// TIA Portal project "Process visualization with HMI" (V15.1)

(* hardware
DEVICE "S71500/ET200MP station_1"  S7-1500 station
   slot 0: "Rail_0"  Rack  6ES7 590-1***0-0AA0
   slot 0: "PM 190W 120/230VAC"  PM 190W 120/230VAC  6EP1333-4BA00
   slot 1: "PLC_1"  CPU 1516-3 PN/DP  6ES7 516-3AN01-0AB0  V2.6
      slot 3: "CPU display_1"  6ES7591-1BA00-0AA0
   slot 2: "DQ 32x24VDC/0.5A HF_1"  DQ 32x24VDC/0.5A HF  6ES7 522-1BL01-0AB0  V1.1
   slot 3: "DI 32x24VDC HF_1"  DI 32x24VDC HF  6ES7 521-1BL00-0AB0  V2.1
   slot 4: "AQ 4xU/I ST_1"  AQ 4xU/I ST  6ES7 532-5HD00-0AB0  V2.2
   slot 5: "AI 8xU/I/RTD/TC ST_1"  AI 8xU/I/RTD/TC ST  6ES7 531-7KF00-0AB0  V2.2
DEVICE "HMI_1"  TP700 Comfort
   slot 0: "HMI_1"  TP700 Comfort  6AV2 124-0GC01-0AX0  15.1.0.0
   slot 1: "HMI_RT_1"  TP700 Comfort  6AV2 124-0GC01-0AX0  15.1.0.0
   slot 5: "HMI_1.IE_CP_1"  PROFINET Interface  15.0.1.0
      slot 1: "PROFINET Interface_1"  PROFINET Interface
         slot 1: "Port_1"  Port
         slot 2: "Port_2"  Port
   slot 7: "HMI_1.MPI/DP_CP_1"  MPI/DP Interface  15.0.1.0
*)

// ===== PLC "PLC_1"  CPU 1516-3 PN/DP =====

VAR_GLOBAL   // PLC tag table "Full_Tag_Table"
   "Panel Emergency Stop" AT %I2.7 : Bool;
   "Start switch" AT %I0.2 : Bool;
   "Stop switch" AT %I0.3 : Bool;
   "Sort area IR" AT %I0.4 : Bool;
   "Sort Area Inductive" AT %I0.5 : Bool;
   "Sort Solenoid Sensor" AT %I0.6 : Bool;
   "Assembly Chute IR" AT %I0.7 : Bool;
   "Assembly Area Through Beam" AT %I1.1 : Bool;
   "Assembly Area Capacitor" AT %I1.2 : Bool;
   "Assembly Area Inductive" AT %I1.3 : Bool;
   "Reject Area IR" AT %I1.4 : Bool;
   "Reject Solenoid Sensor" AT %I1.5 : Bool;
   "Oven Through Beam" AT %I1.6 : Bool;
   "Loading Area Inductive" AT %I1.7 : Bool;
   "Chain Conveyor" AT %Q0.0 : Bool;
   "Sort Solenoid" AT %Q0.1 : Bool;
   "Reject Solenoid" AT %Q0.2 : Bool;
   "Rotary Solenoid" AT %Q0.3 : Bool;
   "Belt Conveyor Direction" AT %Q0.4 : Bool;
   "System Run_Green Lamp" AT %Q3.0 : Bool;
   "Sysyem Stop_Red Lamp" AT %Q3.2 : Bool;
   "Emergency stop" AT %I1.0 : Bool;
   "Ring Queue counter Full" AT %M4.0 : Bool;
   "Sort Solenoid error" AT %M4.3 : Bool;
   "Counter value" AT %MW0 : Int;
   "Reject Solenoid Error" AT %M4.7 : Bool;
   "HMI_Start" AT %M4.1 : Bool;
   "HMI_Stop" AT %M4.2 : Bool;
   "Counter Reset" AT %M4.4 : Bool;
   "DO_card" AT %QD0 : DWord;
   "DI_card" AT %ID0 : DWord;
   "Assembled part counter value" AT %MW4 : Int;
   "HMI_Emergency" AT %M4.5 : Bool;
   "Output metal peg counter value" AT %MW5 : Int;
   "Output plastic ring counter value" AT %MW6 : Int;
   "Input metal peg counter value" AT %MW8 : Int;
   "Input plastic ring counter value" AT %MW10 : Int;
END_VAR

DATA_BLOCK "Conveyors_AUTOMATIC_DB"   // DB1
{ S7_Optimized_Access := 'TRUE' }
VERSION : 0.1
// stored: InstanceOfName Conveyors_AUTOMATIC
"Conveyors_AUTOMATIC"
BEGIN
END_DATA_BLOCK

DATA_BLOCK "Sort Solenoid active_DB"   // DB2
{ S7_Optimized_Access := 'TRUE' }
VERSION : 0.1
// stored: InstanceOfName Sort Solenoid active
"Sort Solenoid active"
BEGIN
END_DATA_BLOCK

DATA_BLOCK "Sort Solenoid active_DB_1"   // DB3
{ S7_Optimized_Access := 'TRUE' }
VERSION : 0.1
// stored: InstanceOfName Sort Solenoid active
"Sort Solenoid active"
BEGIN
END_DATA_BLOCK

DATA_BLOCK "Solenoid Error_DB"   // DB4
{ S7_Optimized_Access := 'TRUE' }
VERSION : 0.1
// stored: InstanceOfName Solenoid Error
"Solenoid Error"
BEGIN
END_DATA_BLOCK

DATA_BLOCK "Counting_DB"   // DB5
{ S7_Optimized_Access := 'TRUE' }
VERSION : 0.1
// stored: InstanceOfName Counter
"Counter"
BEGIN
END_DATA_BLOCK

DATA_BLOCK "Rotary Solenoid1_DB"   // DB6
{ S7_Optimized_Access := 'TRUE' }
VERSION : 0.1
// stored: InstanceOfName Rotary Solenoid1
"Rotary Solenoid1"
BEGIN
END_DATA_BLOCK

DATA_BLOCK "Component Queue Handling_DB"   // DB7
{ S7_Optimized_Access := 'TRUE' }
VERSION : 0.1
// stored: InstanceOfName Component Queue Handling
"Component Queue Handling"
BEGIN
END_DATA_BLOCK

DATA_BLOCK "Solenoid Error_DB_1"   // DB8
{ S7_Optimized_Access := 'TRUE' }
VERSION : 0.1
// stored: InstanceOfName Solenoid Error
"Solenoid Error"
BEGIN
END_DATA_BLOCK

DATA_BLOCK "Assembled part counter_DB"   // DB9
{ S7_Optimized_Access := 'TRUE' }
VERSION : 0.1
// stored: InstanceOfName Assembled part counter
"Assembled part counter"
BEGIN
END_DATA_BLOCK

DATA_BLOCK "Metal peg after assembly counter_DB"   // DB10
{ S7_Optimized_Access := 'TRUE' }
VERSION : 0.1
// stored: InstanceOfName Output metal peg counter
"Output metal peg counter"
BEGIN
END_DATA_BLOCK

DATA_BLOCK "Plastic ring after assembly counter_DB"   // DB11
{ S7_Optimized_Access := 'TRUE' }
VERSION : 0.1
// stored: InstanceOfName Output plastic ring counter
"Output plastic ring counter"
BEGIN
END_DATA_BLOCK

DATA_BLOCK "Input metal peg counter_DB"   // DB12
{ S7_Optimized_Access := 'TRUE' }
VERSION : 0.1
// stored: InstanceOfName Input metal peg counter
"Input metal peg counter"
BEGIN
END_DATA_BLOCK

DATA_BLOCK "Input plastic ring counter_DB"   // DB13
{ S7_Optimized_Access := 'TRUE' }
VERSION : 0.1
// stored: InstanceOfName Input plastic ring counter
"Input plastic ring counter"
BEGIN
END_DATA_BLOCK

FUNCTION_BLOCK "Conveyors_AUTOMATIC"   // FB1, LAD
TITLE = Conveyors Automatic
{ S7_Optimized_Access := 'TRUE' }
VERSION : 0.1
   VAR_INPUT
      "Start Switch" : Bool;
      "Stop Switch" : Bool;
      "Emergency Stop" : Bool;
      "Sort Solenoid Error" : Bool;
      "Panel Emergency Stop" : Bool;
      "Reject Solenoid Error" : Bool;
      H_Start : Bool;
      H_Stop : Bool;
      H_Emergency : Bool;
   END_VAR
   VAR_OUTPUT
      "Chain Conveyor" : Bool;
      "Belt Conveyor" : Bool;
      "System Enable_OK" : Bool;
      "System Enable_not_OK" : Bool;
   END_VAR
   VAR
      Memory_Automatic_Start_Stop : Bool;
   END_VAR
BEGIN

REGION Network 1: System Enable_OK and Conveyor Run
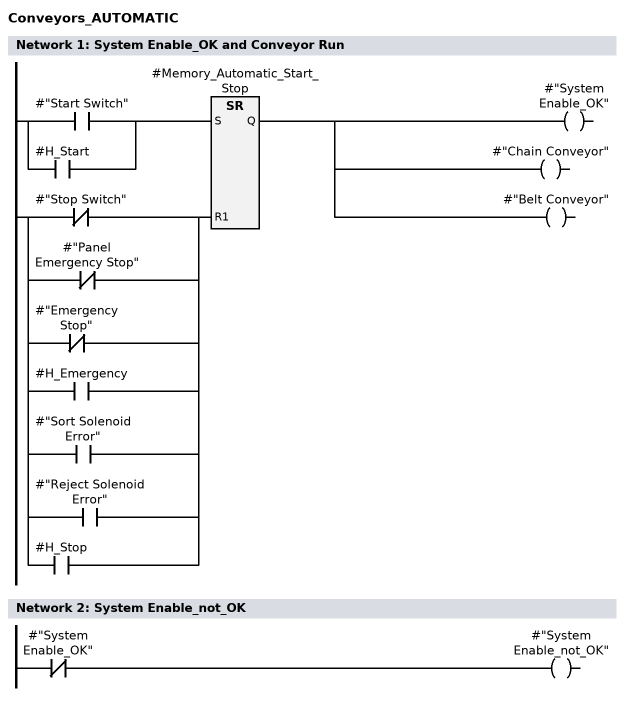
   RUNG wire#powerrail
      Contact( #"Start Switch" )
      wire#w1
      S_SR(operand := #Memory_Automatic_Start_Stop, r1 := wire#w2)
      wire#w3
      Coil( #"System Enable_OK" )
   END_RUNG
   RUNG wire#powerrail
      Contact( #H_Start )
   END_RUNG wire#w1
   RUNG wire#powerrail
      I_Contact( #"Stop Switch" )
   END_RUNG wire#w2
   RUNG wire#powerrail
      I_Contact( #"Panel Emergency Stop" )
   END_RUNG wire#w2
   RUNG wire#powerrail
      I_Contact( #"Emergency Stop" )
   END_RUNG wire#w2
   RUNG wire#powerrail
      Contact( #H_Emergency )
   END_RUNG wire#w2
   RUNG wire#powerrail
      Contact( #"Sort Solenoid Error" )
   END_RUNG wire#w2
   RUNG wire#powerrail
      Contact( #"Reject Solenoid Error" )
   END_RUNG wire#w2
   RUNG wire#powerrail
      Contact( #H_Stop )
   END_RUNG wire#w2
   RUNG wire#w3
      Coil( #"Chain Conveyor" )
   END_RUNG
   RUNG wire#w3
      Coil( #"Belt Conveyor" )
   END_RUNG
   // the same network as SCL:
   IF #"Start Switch" OR #H_Start THEN
       #Memory_Automatic_Start_Stop := TRUE;   // SR flip-flop
   END_IF;
   IF NOT #"Stop Switch" OR NOT #"Panel Emergency Stop" OR NOT #"Emergency Stop" OR #H_Emergency OR #"Sort Solenoid Error" OR #"Reject Solenoid Error" OR #H_Stop THEN
       #Memory_Automatic_Start_Stop := FALSE;
   END_IF;
   #"System Enable_OK" := #Memory_Automatic_Start_Stop;
   #"Chain Conveyor" := #Memory_Automatic_Start_Stop;
   #"Belt Conveyor" := #Memory_Automatic_Start_Stop;
END_REGION

REGION Network 2: System Enable_not_OK
   RUNG wire#powerrail
      I_Contact( #"System Enable_OK" )
      Coil( #"System Enable_not_OK" )
   END_RUNG
   // the same network as SCL:
   #"System Enable_not_OK" := NOT #"System Enable_OK";
END_REGION
END_FUNCTION_BLOCK

FUNCTION_BLOCK "Sort Solenoid active"   // FB2, LAD
TITLE = Sort Solenoid active
{ S7_Optimized_Access := 'TRUE' }
VERSION : 0.1
   VAR_INPUT
      "Sort Area IR" : Bool;
      "Sort Area Inductive" : Bool;
      "Ring Queue counter full" : Bool;
   END_VAR
   VAR_OUTPUT
      "Sort Solenoid" : Bool;
   END_VAR
   VAR
      "Component Pass Delay" : Bool;
      "SR_Sort solenoid on Timer" : Bool;
      "SR_Component pass Delay" : Bool;
      IEC_Timer_0_Instance : TON_TIME;
      IEC_Timer_0_Instance_1 : TON_TIME;
   END_VAR
BEGIN

REGION Network 1: Sort Solenoid activate in case of plastic ring presence
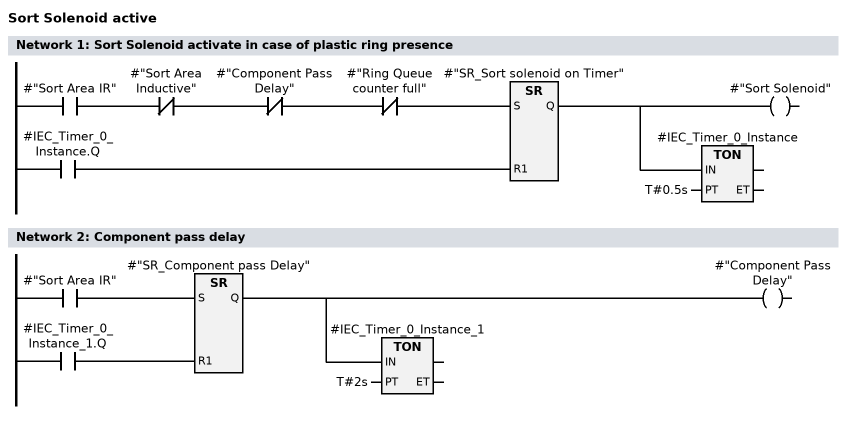
   IF #"Sort Area IR" AND NOT #"Sort Area Inductive" AND NOT #"Component Pass Delay" AND NOT #"Ring Queue counter full" THEN
       #"SR_Sort solenoid on Timer" := TRUE;   // SR flip-flop
   END_IF;
   IF #IEC_Timer_0_Instance.Q THEN #"SR_Sort solenoid on Timer" := FALSE; END_IF;
   #"Sort Solenoid" := #"SR_Sort solenoid on Timer";
   #IEC_Timer_0_Instance(IN := #"SR_Sort solenoid on Timer", PT := T#0.5s);   // TON
END_REGION

REGION Network 2: Component pass delay
   IF #"Sort Area IR" THEN
       #"SR_Component pass Delay" := TRUE;   // SR flip-flop
   END_IF;
   IF #IEC_Timer_0_Instance_1.Q THEN #"SR_Component pass Delay" := FALSE; END_IF;
   #"Component Pass Delay" := #"SR_Component pass Delay";
   #IEC_Timer_0_Instance_1(IN := #"SR_Component pass Delay", PT := T#2s);   // TON
END_REGION
END_FUNCTION_BLOCK

FUNCTION_BLOCK "Solenoid Error"   // FB3, LAD
TITLE = Solenoid error
{ S7_Optimized_Access := 'TRUE' }
VERSION : 0.1
   VAR_INPUT
      "Solenoid on" : Bool;
      "Solenoid sensor" : Bool;
   END_VAR
   VAR_OUTPUT
      "Solenoid error" : Bool;
   END_VAR
   VAR
      "Hold off delay" : Bool;
      IEC_Timer_0_Instance : TON_TIME;
   END_VAR
BEGIN

REGION Network 1: Solenoid error
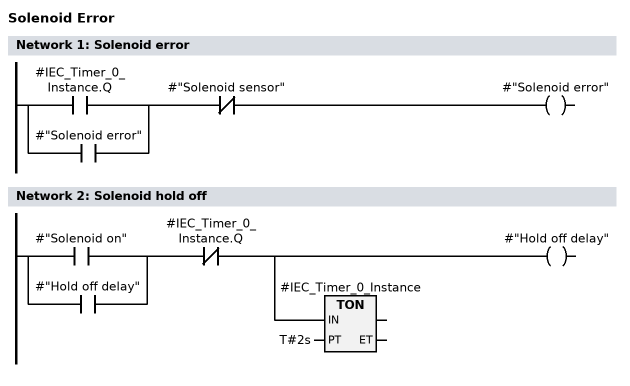
   RUNG wire#powerrail
      Contact( #IEC_Timer_0_Instance.Q )
      wire#w1
      I_Contact( #"Solenoid sensor" )
      Coil( #"Solenoid error" )
   END_RUNG
   RUNG wire#powerrail
      Contact( #"Solenoid error" )
   END_RUNG wire#w1
   // the same network as SCL:
   #"Solenoid error" := (#IEC_Timer_0_Instance.Q OR #"Solenoid error") AND NOT #"Solenoid sensor";
END_REGION

REGION Network 2: Solenoid hold off
   #"Hold off delay" := (#"Solenoid on" OR #"Hold off delay") AND NOT #IEC_Timer_0_Instance.Q;
   #IEC_Timer_0_Instance(IN := #"Hold off delay", PT := T#2s);   // TON
END_REGION
END_FUNCTION_BLOCK

FUNCTION_BLOCK "Counter"   // FB4, LAD
{ S7_Optimized_Access := 'TRUE' }
VERSION : 0.1
   VAR_INPUT
      "Sort Solenoid" : Bool;
      "Rotary Solenoid" : Bool;
      "Reset counter" : Bool;
   END_VAR
   VAR_OUTPUT
      "Counter value" : Int;
      "Ring Queue counter full" : Bool;
   END_VAR
   VAR RETAIN
      IEC_Counter_0_Instance : CTUD_INT;
   END_VAR
BEGIN

REGION Network 1
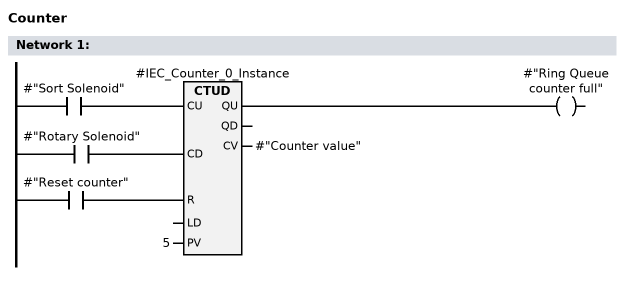
   #IEC_Counter_0_Instance(CU := #"Sort Solenoid",   // CTUD
                           CD := #"Rotary Solenoid",
                           R := #"Reset counter",
                           PV := 5,
                           CV => #"Counter value");
   #"Ring Queue counter full" := #IEC_Counter_0_Instance.QU;
END_REGION
END_FUNCTION_BLOCK

FUNCTION_BLOCK "Rotary Solenoid1"   // FB5, LAD
{ S7_Optimized_Access := 'TRUE' }
VERSION : 0.1
   VAR_INPUT
      "Assembly chute IR" : Bool;
      "Counter value" : Int;
   END_VAR
   VAR_OUTPUT
      "Rotary Solenoid" : Bool;
   END_VAR
   VAR
      "Rotary Solenoid on Timer" : Bool;
      IEC_Timer_0_Instance : TON_TIME;
      "Component pass delay" : Bool;
      "SR_Component pass delay" : Bool;
      IEC_Timer_0_Instance_2 : TON_TIME;
      IEC_Timer_0_Instance_1 : TON_TIME;
   END_VAR
BEGIN

REGION Network 1: Rotary Solenoid
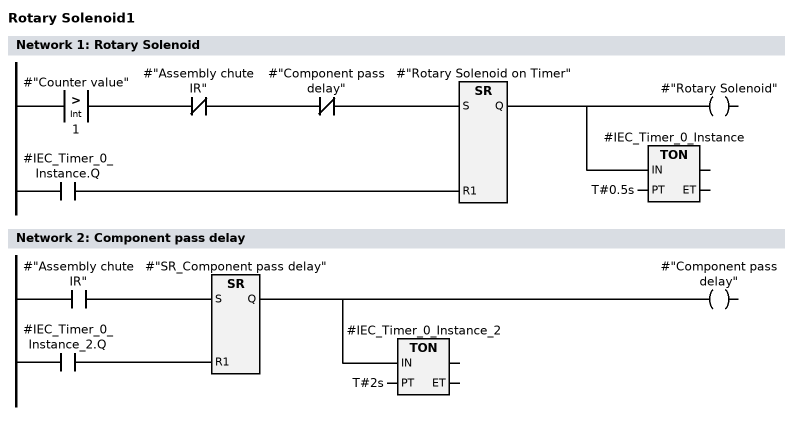
   IF (#"Counter value" > 1) AND NOT #"Assembly chute IR" AND NOT #"Component pass delay" THEN
       #"Rotary Solenoid on Timer" := TRUE;   // SR flip-flop
   END_IF;
   IF #IEC_Timer_0_Instance.Q THEN #"Rotary Solenoid on Timer" := FALSE; END_IF;
   #"Rotary Solenoid" := #"Rotary Solenoid on Timer";
   #IEC_Timer_0_Instance(IN := #"Rotary Solenoid on Timer", PT := T#0.5s);   // TON
END_REGION

REGION Network 2: Component pass delay
   IF #"Assembly chute IR" THEN
       #"SR_Component pass delay" := TRUE;   // SR flip-flop
   END_IF;
   IF #IEC_Timer_0_Instance_2.Q THEN #"SR_Component pass delay" := FALSE; END_IF;
   #"Component pass delay" := #"SR_Component pass delay";
   #IEC_Timer_0_Instance_2(IN := #"SR_Component pass delay", PT := T#2s);   // TON
END_REGION
END_FUNCTION_BLOCK

FUNCTION_BLOCK "Component Queue Handling"   // FB6, LAD
TITLE = Component Queue Handling
{ S7_Optimized_Access := 'TRUE' }
VERSION : 0.1
   VAR_INPUT
      "Start Switch" : Bool;
      "Assembly Area Capacitive" : Bool;
      "Assembly Area Inductive" : Bool;
      "Reject Area IR" : Bool;
      "Assembly Area Through Beam" : Bool;
   END_VAR
   VAR_OUTPUT
      "Reject Solenoid" : Bool;
   END_VAR
   VAR
      "Assembly Complete" : Bool;
      "Pointer Register" : Word;
      "Data Register" : Word;
      "SHL Memory" : Bool;
      "SHR Memory" : Bool;
      "And Result" : Word;
      SR_Reject : Bool;
      IEC_Timer_0_Instance : TON_TIME;
   END_VAR
   VAR_TEMP   // added for the SCL form of the ladder/FBD networks
      _w1 : Bool;
   END_VAR
BEGIN

REGION Network 1: data and pointer register
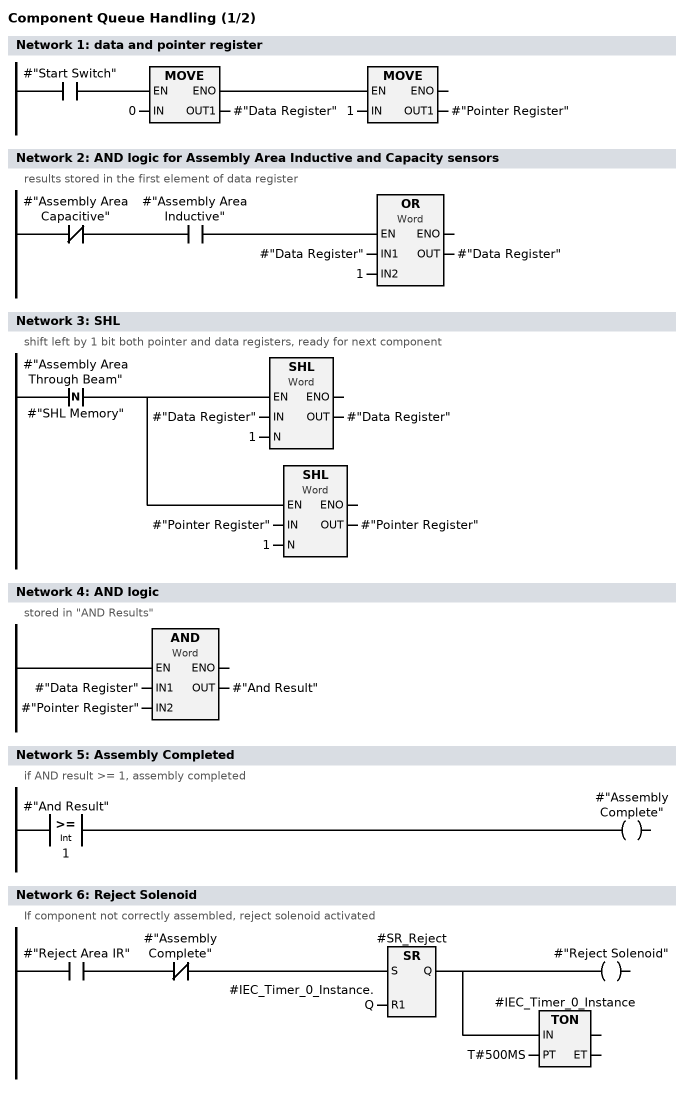
   RUNG wire#powerrail
      Contact( #"Start Switch" )
      Move(in := 0, out1 => #"Data Register")
      Move(in := 1, out1 => #"Pointer Register")
   END_RUNG
   // the same network as SCL:
   IF #"Start Switch" THEN
       #"Data Register" := 0;
       #"Pointer Register" := 1;
   END_IF;
END_REGION

REGION Network 2: AND logic for Assembly Area Inductive and Capacity sensors
   // results stored in the first element of data register
   IF NOT #"Assembly Area Capacitive" AND #"Assembly Area Inductive" THEN
       #"Data Register" := #"Data Register" OR 1;
   END_IF;
END_REGION

REGION Network 3: SHL
   // shift left by 1 bit both pointer and data registers, ready for next component
   RUNG wire#powerrail
      N_Contact(operand := #"Assembly Area Through Beam", bit := #"SHL Memory")
      wire#w1
      { S7_Templates := "SrcType := Word" } Shl(in := #"Data Register", n := 1, out => #"Data Register")
   END_RUNG
   RUNG wire#w1
      { S7_Templates := "SrcType := Word" } Shl(in := #"Pointer Register", n := 1, out => #"Pointer Register")
   END_RUNG
   // the same network as SCL:
   #_w1 := NOT #"Assembly Area Through Beam" AND #"SHL Memory";   // falling edge of #"Assembly Area Through Beam"
   #"SHL Memory" := #"Assembly Area Through Beam";
   IF #_w1 THEN
       #"Data Register" := SHL(IN := #"Data Register", N := 1);
       #"Pointer Register" := SHL(IN := #"Pointer Register", N := 1);
   END_IF;
END_REGION

REGION Network 4: AND logic
   // stored in "AND Results"
   RUNG wire#powerrail
      { S7_Templates := "SrcType := Word" } And(in1 := #"Data Register", in2 := #"Pointer Register", out => #"And Result")
   END_RUNG
   // the same network as SCL:
   #"And Result" := #"Data Register" AND #"Pointer Register";
END_REGION

REGION Network 5: Assembly Completed
   // if AND result >= 1, assembly completed
   RUNG wire#powerrail
      { S7_Templates := "SrcType := Int" } GE_Contact(in1 := #"And Result", in2 := 1)
      Coil( #"Assembly Complete" )
   END_RUNG
   // the same network as SCL:
   #"Assembly Complete" := #"And Result" >= 1;
END_REGION

REGION Network 6: Reject Solenoid
   // If component not correctly assembled, reject solenoid activated
   IF #"Reject Area IR" AND NOT #"Assembly Complete" THEN
       #SR_Reject := TRUE;   // SR flip-flop
   END_IF;
   IF #IEC_Timer_0_Instance.Q THEN #SR_Reject := FALSE; END_IF;
   #"Reject Solenoid" := #SR_Reject;
   #IEC_Timer_0_Instance(IN := #SR_Reject, PT := T#500MS);   // TON
END_REGION

REGION Network 7: SHR
   // when component left assembly area, shift right by 1 bit
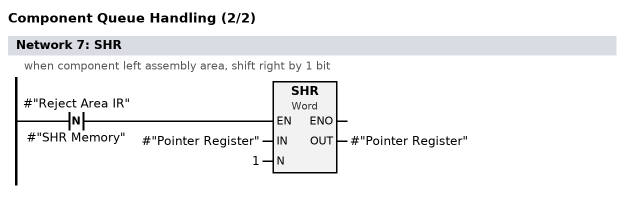
   RUNG wire#powerrail
      N_Contact(operand := #"Reject Area IR", bit := #"SHR Memory")
      { S7_Templates := "SrcType := Word" } Shr(in := #"Pointer Register", n := 1, out => #"Pointer Register")
   END_RUNG
   // the same network as SCL:
   #_w1 := NOT #"Reject Area IR" AND #"SHR Memory";   // falling edge of #"Reject Area IR"
   #"SHR Memory" := #"Reject Area IR";
   IF #_w1 THEN #"Pointer Register" := SHR(IN := #"Pointer Register", N := 1); END_IF;
END_REGION
END_FUNCTION_BLOCK

FUNCTION_BLOCK "Assembled part counter"   // FB7, LAD
TITLE = Assembled part counter
{ S7_Optimized_Access := 'TRUE' }
VERSION : 0.1
   VAR_INPUT
      "Reject area IR" : Bool;
      "Reject solenoid" : Bool;
      "Reset counter" : Bool;
   END_VAR
   VAR_OUTPUT
      "Assembled part counter value" : Int;
   END_VAR
   VAR RETAIN
      IEC_Counter_0_Instance : CTU_INT;
   END_VAR
BEGIN

REGION Network 1: Counter for assembled parts
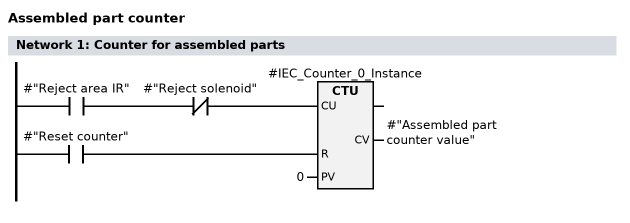
   #IEC_Counter_0_Instance(CU := #"Reject area IR" AND NOT #"Reject solenoid",   // CTU
                           R := #"Reset counter",
                           PV := 0,
                           CV => #"Assembled part counter value");
END_REGION
END_FUNCTION_BLOCK

FUNCTION_BLOCK "Output metal peg counter"   // FB8, LAD
{ S7_Optimized_Access := 'TRUE' }
VERSION : 0.1
   VAR_INPUT
      "Assembly Area Inductive" : Bool;
      "Assembly Area Capacitive" : Bool;
      "Assembly Area thru beam" : Bool;
      "Reset counter" : Bool;
   END_VAR
   VAR_OUTPUT
      "Metal peg" : Int;
   END_VAR
   VAR RETAIN
      IEC_Counter_0_Instance : CTU_INT;
   END_VAR
BEGIN

REGION Network 1: Metal peg counter
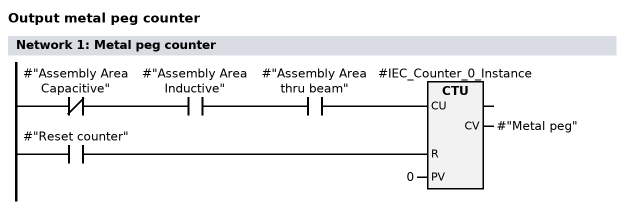
   #IEC_Counter_0_Instance(CU := NOT #"Assembly Area Capacitive" AND #"Assembly Area Inductive" AND #"Assembly Area thru beam",   // CTU
                           R := #"Reset counter",
                           PV := 0,
                           CV => #"Metal peg");
END_REGION
END_FUNCTION_BLOCK

FUNCTION_BLOCK "Output plastic ring counter"   // FB9, LAD
{ S7_Optimized_Access := 'TRUE' }
VERSION : 0.1
   VAR_INPUT
      "Assembly Area Inductive" : Bool;
      "Assembly Area Capacitive" : Bool;
      "Assembly Area thru beam" : Bool;
      "Reset counter" : Bool;
   END_VAR
   VAR_OUTPUT
      "Plastic ring" : Int;
   END_VAR
   VAR RETAIN
      IEC_Counter_0_Instance : CTU_INT;
   END_VAR
BEGIN

REGION Network 1: Plastic ring counter
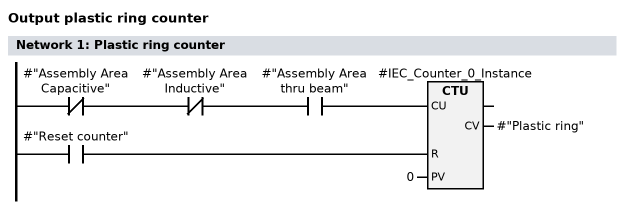
   #IEC_Counter_0_Instance(CU := NOT #"Assembly Area Capacitive" AND NOT #"Assembly Area Inductive" AND #"Assembly Area thru beam",   // CTU
                           R := #"Reset counter",
                           PV := 0,
                           CV => #"Plastic ring");
END_REGION
END_FUNCTION_BLOCK

FUNCTION_BLOCK "Input metal peg counter"   // FB10, LAD
{ S7_Optimized_Access := 'TRUE' }
VERSION : 0.1
   VAR_INPUT
      "Sort Area IR" : Bool;
      "Sort Area inductive" : Bool;
      "Reset counter" : Bool;
   END_VAR
   VAR_OUTPUT
      "Input metal peg" : Int;
   END_VAR
   VAR RETAIN
      IEC_Counter_0_Instance : CTU_INT;
   END_VAR
BEGIN

REGION Network 1: Input Metal Peg counter
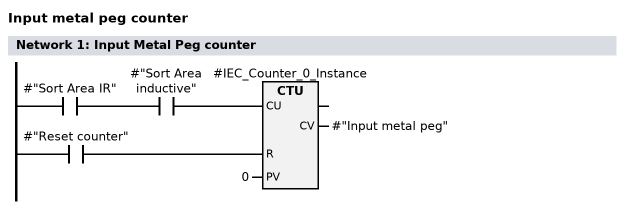
   #IEC_Counter_0_Instance(CU := #"Sort Area IR" AND #"Sort Area inductive",   // CTU
                           R := #"Reset counter",
                           PV := 0,
                           CV => #"Input metal peg");
END_REGION
END_FUNCTION_BLOCK

FUNCTION_BLOCK "Input plastic ring counter"   // FB11, LAD
{ S7_Optimized_Access := 'TRUE' }
VERSION : 0.1
   VAR_INPUT
      "Sort Area IR" : Bool;
      "Sort Area inductive" : Bool;
      "Reset counter" : Bool;
   END_VAR
   VAR_OUTPUT
      "Input plastic ring" : Int;
   END_VAR
   VAR RETAIN
      IEC_Counter_0_Instance : CTU_INT;
   END_VAR
BEGIN

REGION Network 1: Input plastic ring counter
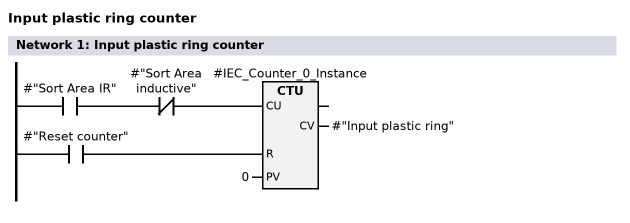
   #IEC_Counter_0_Instance(CU := #"Sort Area IR" AND NOT #"Sort Area inductive",   // CTU
                           R := #"Reset counter",
                           PV := 0,
                           CV => #"Input plastic ring");
END_REGION
END_FUNCTION_BLOCK

ORGANIZATION_BLOCK "Main"   // OB1, LAD, ProgramCycle
TITLE = "Main Program Sweep (Cycle)"
{ S7_Optimized_Access := 'TRUE' }
VERSION : 0.1
   VAR_INPUT
      Initial_Call : Bool;   // Initial call of this OB
      Remanence : Bool;   // =True, if remanent data are available
   END_VAR
BEGIN

REGION Network 1: System Run OK and conveyors start
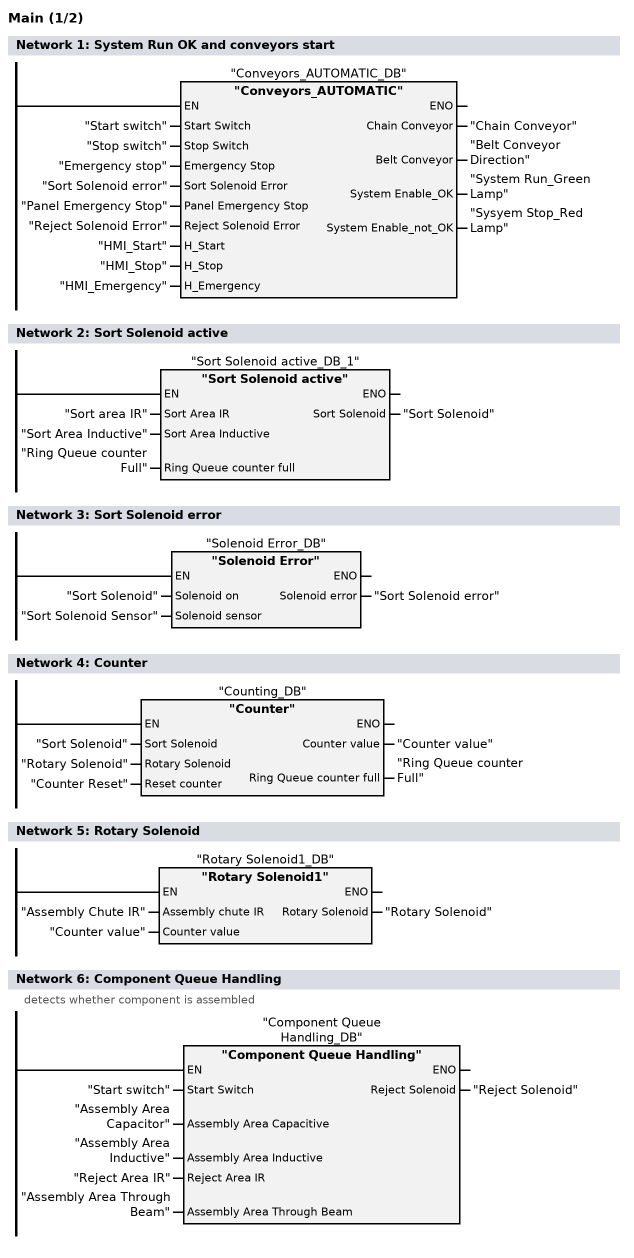
   RUNG wire#powerrail
      "Conveyors_AUTOMATIC_DB"("Start Switch" := "Start switch", "Stop Switch" := "Stop switch", "Emergency Stop" := "Emergency stop", "Sort Solenoid Error" := "Sort Solenoid error", "Panel Emergency Stop" := "Panel Emergency Stop", "Reject Solenoid Error" := "Reject Solenoid Error", H_Start := "HMI_Start", H_Stop := "HMI_Stop", H_Emergency := "HMI_Emergency", "Chain Conveyor" => "Chain Conveyor", "Belt Conveyor" => "Belt Conveyor Direction", "System Enable_OK" => "System Run_Green Lamp", "System Enable_not_OK" => "Sysyem Stop_Red Lamp")
   END_RUNG
   // the same network as SCL:
   "Conveyors_AUTOMATIC_DB"("Start Switch" := "Start switch",   // "Conveyors_AUTOMATIC"
                           "Stop Switch" := "Stop switch",
                           "Emergency Stop" := "Emergency stop",
                           "Sort Solenoid Error" := "Sort Solenoid error",
                           "Panel Emergency Stop" := "Panel Emergency Stop",
                           "Reject Solenoid Error" := "Reject Solenoid Error",
                           H_Start := "HMI_Start",
                           H_Stop := "HMI_Stop",
                           H_Emergency := "HMI_Emergency",
                           "Chain Conveyor" => "Chain Conveyor",
                           "Belt Conveyor" => "Belt Conveyor Direction",
                           "System Enable_OK" => "System Run_Green Lamp",
                           "System Enable_not_OK" => "Sysyem Stop_Red Lamp");
END_REGION

REGION Network 2: Sort Solenoid active
   RUNG wire#powerrail
      "Sort Solenoid active_DB_1"("Sort Area IR" := "Sort area IR", "Sort Area Inductive" := "Sort Area Inductive", "Ring Queue counter full" := "Ring Queue counter Full", "Sort Solenoid" => "Sort Solenoid")
   END_RUNG
   // the same network as SCL:
   "Sort Solenoid active_DB_1"("Sort Area IR" := "Sort area IR",   // "Sort Solenoid active"
                           "Sort Area Inductive" := "Sort Area Inductive",
                           "Ring Queue counter full" := "Ring Queue counter Full",
                           "Sort Solenoid" => "Sort Solenoid");
END_REGION

REGION Network 3: Sort Solenoid error
   RUNG wire#powerrail
      "Solenoid Error_DB"("Solenoid on" := "Sort Solenoid", "Solenoid sensor" := "Sort Solenoid Sensor", "Solenoid error" => "Sort Solenoid error")
   END_RUNG
   // the same network as SCL:
   "Solenoid Error_DB"("Solenoid on" := "Sort Solenoid",   // "Solenoid Error"
                       "Solenoid sensor" := "Sort Solenoid Sensor",
                       "Solenoid error" => "Sort Solenoid error");
END_REGION

REGION Network 4: Counter
   RUNG wire#powerrail
      "Counting_DB"("Sort Solenoid" := "Sort Solenoid", "Rotary Solenoid" := "Rotary Solenoid", "Reset counter" := "Counter Reset", "Counter value" => "Counter value", "Ring Queue counter full" => "Ring Queue counter Full")
   END_RUNG
   // the same network as SCL:
   "Counting_DB"("Sort Solenoid" := "Sort Solenoid",   // "Counter"
                 "Rotary Solenoid" := "Rotary Solenoid",
                 "Reset counter" := "Counter Reset",
                 "Counter value" => "Counter value",
                 "Ring Queue counter full" => "Ring Queue counter Full");
END_REGION

REGION Network 5: Rotary Solenoid
   RUNG wire#powerrail
      "Rotary Solenoid1_DB"("Assembly chute IR" := "Assembly Chute IR", "Counter value" := "Counter value", "Rotary Solenoid" => "Rotary Solenoid")
   END_RUNG
   // the same network as SCL:
   "Rotary Solenoid1_DB"("Assembly chute IR" := "Assembly Chute IR",   // "Rotary Solenoid1"
                         "Counter value" := "Counter value",
                         "Rotary Solenoid" => "Rotary Solenoid");
END_REGION

REGION Network 6: Component Queue Handling
   // detects whether component is assembled
   RUNG wire#powerrail
      "Component Queue Handling_DB"("Start Switch" := "Start switch", "Assembly Area Capacitive" := "Assembly Area Capacitor", "Assembly Area Inductive" := "Assembly Area Inductive", "Reject Area IR" := "Reject Area IR", "Assembly Area Through Beam" := "Assembly Area Through Beam", "Reject Solenoid" => "Reject Solenoid")
   END_RUNG
   // the same network as SCL:
   "Component Queue Handling_DB"("Start Switch" := "Start switch",   // "Component Queue Handling"
                           "Assembly Area Capacitive" := "Assembly Area Capacitor",
                           "Assembly Area Inductive" := "Assembly Area Inductive",
                           "Reject Area IR" := "Reject Area IR",
                           "Assembly Area Through Beam" := "Assembly Area Through Beam",
                           "Reject Solenoid" => "Reject Solenoid");
END_REGION

REGION Network 7: Reject Solenoid error
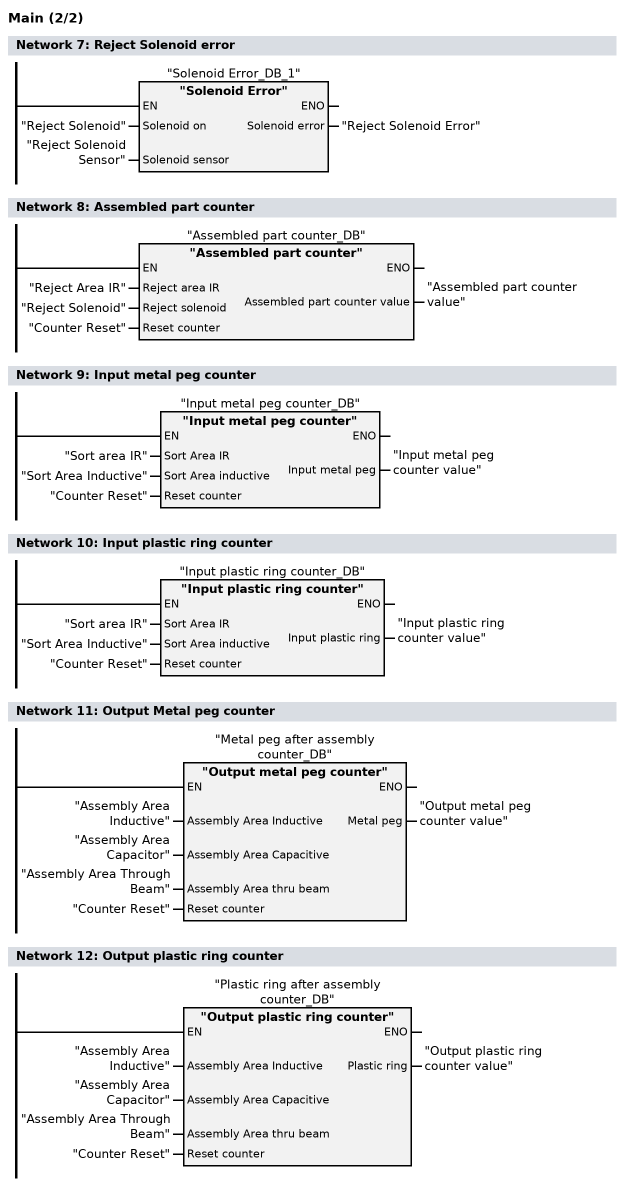
   RUNG wire#powerrail
      "Solenoid Error_DB_1"("Solenoid on" := "Reject Solenoid", "Solenoid sensor" := "Reject Solenoid Sensor", "Solenoid error" => "Reject Solenoid Error")
   END_RUNG
   // the same network as SCL:
   "Solenoid Error_DB_1"("Solenoid on" := "Reject Solenoid",   // "Solenoid Error"
                         "Solenoid sensor" := "Reject Solenoid Sensor",
                         "Solenoid error" => "Reject Solenoid Error");
END_REGION

REGION Network 8: Assembled part counter
   RUNG wire#powerrail
      "Assembled part counter_DB"("Reject area IR" := "Reject Area IR", "Reject solenoid" := "Reject Solenoid", "Reset counter" := "Counter Reset", "Assembled part counter value" => "Assembled part counter value")
   END_RUNG
   // the same network as SCL:
   "Assembled part counter_DB"("Reject area IR" := "Reject Area IR",   // "Assembled part counter"
                           "Reject solenoid" := "Reject Solenoid",
                           "Reset counter" := "Counter Reset",
                           "Assembled part counter value" => "Assembled part counter value");
END_REGION

REGION Network 9: Input metal peg counter
   RUNG wire#powerrail
      "Input metal peg counter_DB"("Sort Area IR" := "Sort area IR", "Sort Area inductive" := "Sort Area Inductive", "Reset counter" := "Counter Reset", "Input metal peg" => "Input metal peg counter value")
   END_RUNG
   // the same network as SCL:
   "Input metal peg counter_DB"("Sort Area IR" := "Sort area IR",   // "Input metal peg counter"
                           "Sort Area inductive" := "Sort Area Inductive",
                           "Reset counter" := "Counter Reset",
                           "Input metal peg" => "Input metal peg counter value");
END_REGION

REGION Network 10: Input plastic ring counter
   RUNG wire#powerrail
      "Input plastic ring counter_DB"("Sort Area IR" := "Sort area IR", "Sort Area inductive" := "Sort Area Inductive", "Reset counter" := "Counter Reset", "Input plastic ring" => "Input plastic ring counter value")
   END_RUNG
   // the same network as SCL:
   "Input plastic ring counter_DB"("Sort Area IR" := "Sort area IR",   // "Input plastic ring counter"
                           "Sort Area inductive" := "Sort Area Inductive",
                           "Reset counter" := "Counter Reset",
                           "Input plastic ring" => "Input plastic ring counter value");
END_REGION

REGION Network 11: Output Metal peg counter
   RUNG wire#powerrail
      "Metal peg after assembly counter_DB"("Assembly Area Inductive" := "Assembly Area Inductive", "Assembly Area Capacitive" := "Assembly Area Capacitor", "Assembly Area thru beam" := "Assembly Area Through Beam", "Reset counter" := "Counter Reset", "Metal peg" => "Output metal peg counter value")
   END_RUNG
   // the same network as SCL:
   "Metal peg after assembly counter_DB"("Assembly Area Inductive" := "Assembly Area Inductive",   // "Output metal peg counter"
                           "Assembly Area Capacitive" := "Assembly Area Capacitor",
                           "Assembly Area thru beam" := "Assembly Area Through Beam",
                           "Reset counter" := "Counter Reset",
                           "Metal peg" => "Output metal peg counter value");
END_REGION

REGION Network 12: Output plastic ring counter
   RUNG wire#powerrail
      "Plastic ring after assembly counter_DB"("Assembly Area Inductive" := "Assembly Area Inductive", "Assembly Area Capacitive" := "Assembly Area Capacitor", "Assembly Area thru beam" := "Assembly Area Through Beam", "Reset counter" := "Counter Reset", "Plastic ring" => "Output plastic ring counter value")
   END_RUNG
   // the same network as SCL:
   "Plastic ring after assembly counter_DB"("Assembly Area Inductive" := "Assembly Area Inductive",   // "Output plastic ring counter"
                           "Assembly Area Capacitive" := "Assembly Area Capacitor",
                           "Assembly Area thru beam" := "Assembly Area Through Beam",
                           "Reset counter" := "Counter Reset",
                           "Plastic ring" => "Output plastic ring counter value");
END_REGION
END_ORGANIZATION_BLOCK

(* ===== HMI "HMI_RT_1" =====
system functions are stored by id; their names below are inferred from use
connection "HMI_Connection_1": ETHERNET, S7_1500_OMS

HMI tags "Default tag table"
   "Counter value" : Int = PLC "Counter value" AT %MW0, 100 ms
   "Sort Solenoid Sensor" : Bool = PLC "Sort Solenoid Sensor" AT %I0.6, 100 ms
   "Ring Queue counter Full" : Bool = PLC "Ring Queue counter Full" AT %M4.0, 100 ms
   "Counter Reset" : Bool = PLC "Counter Reset" AT %M4.4, 100 ms
   "HMI_Stop" : Bool = PLC HMI_Stop AT %M4.2, 100 ms
   "HMI_Start" : Bool = PLC HMI_Start AT %M4.1, 100 ms
   "Emergency stop" : Bool = PLC "Emergency stop" AT %I1.0, 100 ms
   "Stop switch" : Bool = PLC "Stop switch" AT %I0.3, 100 ms
   "System Run_Green Lamp" : Bool = PLC "System Run_Green Lamp" AT %Q3.0, 100 ms
   "Sysyem Stop_Red Lamp" : Bool = PLC "Sysyem Stop_Red Lamp" AT %Q3.2, 100 ms
   "Chain Conveyor" : Bool = PLC "Chain Conveyor" AT %Q0.0, 100 ms
   "Sort area IR" : Bool = PLC "Sort area IR" AT %I0.4, 100 ms
   "Sort Area Inductive" : Bool = PLC "Sort Area Inductive" AT %I0.5, 100 ms
   "Assembly Area Inductive" : Bool = PLC "Assembly Area Inductive" AT %I1.3, 100 ms
   "Assembly Area Capacitor" : Bool = PLC "Assembly Area Capacitor" AT %I1.2, 100 ms
   "Assembly Chute IR" : Bool = PLC "Assembly Chute IR" AT %I0.7, 100 ms
   "Reject Solenoid" : Bool = PLC "Reject Solenoid" AT %Q0.2, 100 ms
   "Reject Solenoid Sensor" : Bool = PLC "Reject Solenoid Sensor" AT %I1.5, 100 ms
   "Belt Conveyor Direction" : Bool = PLC "Belt Conveyor Direction" AT %Q0.4, 100 ms
   "Assembly Area Through Beam" : Bool = PLC "Assembly Area Through Beam" AT %I1.1, 100 ms
   "Assembled part counter value" : Int = PLC "Assembled part counter value" AT %MW4, 100 ms
   "HMI_Emergency" : Bool = PLC HMI_Emergency AT %M4.5, 100 ms
   "Metal peg counter value" : Int = PLC "Output metal peg counter value" AT %MW5, 1 s
   "Plastic ring counter value" : Int = PLC "Output plastic ring counter value" AT %MW6, 1 s
   "Input metal peg counter value" : Int = PLC "Input metal peg counter value" AT %MW8, 1 s
   "Input plastic ring counter value" : Int = PLC "Input plastic ring counter value" AT %MW10, 1 s

Template "Template_1" 800x480
   Button "Exit" at 720,420 size 78x58; TextOff 'Exit'; PictureOff "ExitRuntime_TP700_Comfort_TR"; PictureOn "ExitRuntime_TP700_Comfort_TR"
      on Release: StopRuntime(0)
   Button "Template_Button" at 640,420 size 78x58; TextOff 'Text'
   Button "Template_Button_1" at 560,420 size 78x58; TextOff 'Text'
   Button "Template_Button_2" at 480,420 size 78x58; TextOff 'Text'
   Button "Template_Button_3" at 400,420 size 78x58; TextOff 'Text'
   Button "Template_Button_4" at 321,420 size 78x58; TextOff 'Text'
   Button "Template_Button_5" at 241,420 size 78x58; TextOff 'Text'
   Button "Template_Button_6" at 161,420 size 78x58; TextOff 'Text'
   Button "Template_Button_7" at 81,420 size 78x58; TextOff 'Text'
   Button "Start screen" at 1,420 size 78x58; TextOff 'Start screen'; PictureOff "NavigateHome_TP700_Comfort_TR"; PictureOn "NavigateHome_TP700_Comfort_TR"
      on Release: ActivateScreen("Sorting Station Overview", 0)

screen "Sorting Station Overview" 800x480, template "Template_1"
   TextField "HmiScreenItemData_5" at 80,196 size 640x25; Text 'Welcome to HMI_1 (TP700 Comfort)!'
   Button "HmiScreenItemData" at 36,36 size 159x47; TextOff 'System Control'; PictureOff "Navigates to System Control for TP700 Comfort 15.1.0.0"; PictureOn "Navigates to System Control for TP700 Comfort 15.1.0.0"
      on Release: ActivateScreen("System Control", 0)
   Button "HmiScreenItemData_1" at 36,95 size 159x47; TextOff 'Input/Output'; PictureOff "Navigates to Input/Output for TP700 Comfort 15.1.0.0"; PictureOn "Navigates to Input/Output for TP700 Comfort 15.1.0.0"
      on Release: ActivateScreen("Input/Output", 0)
   Button "HmiScreenItemData_2" at 36,154 size 159x47; TextOff 'Temperature Control'; PictureOff "Navigates to Temperature Control for TP700 Comfort 15.1.0.0"; PictureOn "Navigates to Temperature Control for TP700 Comfort 15.1.0.0"
      on Release: ActivateScreen("Temperature Control", 0)
   Button "HmiScreenItemData_3" at 36,213 size 159x47; TextOff 'Alarm'; PictureOff "Navigates to Alarm for TP700 Comfort 15.1.0.0"; PictureOn "Navigates to Alarm for TP700 Comfort 15.1.0.0"
      on Release: ActivateScreen("Alarm", 0)
   Button "HmiScreenItemData_4" at 36,272 size 159x47; TextOff 'Exercise'; PictureOff "Navigates to Exercise for TP700 Comfort 15.1.0.0"; PictureOn "Navigates to Exercise for TP700 Comfort 15.1.0.0"
      on Release: ActivateScreen("Exercise", 0)
   Button "HmiScreenItemData_6" at 36,331 size 159x47; TextOff 'System screens'; PictureOff "Navigates to System screens for TP700 Comfort 15.1.0.0"; PictureOn "Navigates to System screens for TP700 Comfort 15.1.0.0"
      on Release: ActivateScreen("System screens", 0)
   GraphicView "Graphic view_1" at 230,64 size 473x289; Picture "HMI picture"

screen "System Control" 800x480, template "Template_1"
   Button "Back" at 1,1 size 159x47; TextOff 'Back'
      on Release: ActivateScreen("Sorting Station Overview", 0)
   GraphicView "Graphic view_1" at 0,0 size 800x480; Picture "bytronic"
   Button "Back_1" at 0,28 size 159x47; TextOn 'Back'; TextOff 'Back'
      on Release: ActivateScreen("Sorting Station Overview", 0)
   IOField "I/O field_1" at 23,335 size 29x32; FormatPattern 9
      ProcessValue <- "Counter value"
   TextField "Text field_1" at 7,283 size 134x23; Text 'Counter Value'
   Circle "Circle_1" at 241,32 size 18x18
      Appearance <- "Sort Solenoid Sensor"
   Circle "Circle_2" at 65,331 size 35x35
      Appearance <- "Ring Queue counter Full"
   Button "Button_1" at 283,412 size 40x40; TextOff 'Text'; PictureOn "Pushbutton_Round_R_On_256c"; PictureOff "Pushbutton_Round_R_Off_256c"
      on Press: function_b14e0dd5("Counter Reset", 0)
   Button "Button_2" at 139,412 size 40x40; TextOff 'Text'; PictureOn "Pushbutton_Round_R_On_256c"; PictureOff "Pushbutton_Round_R_Off_256c"
      on Press: function_b14e0dd5("HMI_Stop", 0)
   Button "Button_3" at 182,412 size 40x40; TextOff 'Text'; PictureOn "Pushbutton_Round_G_On_256c"; PictureOff "Pushbutton_Round_G_Off_256c"
      on Press: function_b14e0dd5("HMI_Start", 0)
   Circle "Circle_3" at 240,108 size 20x20
      Appearance <- "Sort Area Inductive"
   Circle "Circle_4" at 418,387 size 25x25
      Appearance <- "Sysyem Stop_Red Lamp"
   Circle "Circle_5" at 418,413 size 25x25
      Appearance <- "Emergency stop"
   Circle "Circle_6" at 418,439 size 25x25
      Appearance <- "System Run_Green Lamp"
   Rectangle "Rectangle_1" at 131,153 size 28x18
      Appearance <- "Chain Conveyor"
   Rectangle "Rectangle_2" at 224,101 size 9x24
      Appearance <- "Sort area IR"
   Rectangle "Rectangle_3" at 308,218 size 27x19
      Appearance <- "Assembly Area Capacitor"
   Circle "Circle_7" at 313,275 size 18x18
      Appearance <- "Assembly Area Inductive"
   Rectangle "Rectangle_4" at 241,295 size 18x10
      Appearance <- "Assembly Chute IR"
   Circle "Circle_8" at 498,347 size 16x16
      Appearance <- "Reject Solenoid Sensor"
   Rectangle "Rectangle_5" at 519,334 size 19x25
      Appearance <- "Belt Conveyor Direction"
   Circle "Circle_9" at 343,253 size 14x14
      Appearance <- "Assembly Area Through Beam"
   IOField "I/O field_2" at 728,378 size 63x25; FormatPattern 999
      ProcessValue <- "Assembled part counter value"
   Switch "Switch_1" at 1,378 size 100x100; CaptionText 'Switch'; TextOff 'OFF'; TextOn 'ON'; PictureOn "Pushbutton_Emergency_On_256c"; PictureOff "Pushbutton_Emergency_Off_256c"
      on SwitchOn: SetBit("HMI_Emergency")
   IOField "I/O field_3" at 653,378 size 63x25; FormatPattern 999
      ProcessValue <- "Metal peg counter value"
   IOField "I/O field_4" at 576,378 size 63x25; FormatPattern 999
      ProcessValue <- "Plastic ring counter value"

screen "Input/Output" 800x480, template "Template_1"
   Button "Back" at 1,1 size 159x47; TextOff 'Back'
      on Release: ActivateScreen("Sorting Station Overview", 0)
   TextField "Text field_1" at 43,63 size 134x23; Text 'Counter Value'
   TextField "Text field_2" at 269,62 size 63x23; Text 'Inputs'
   TextField "Text field_3" at 545,63 size 76x23; Text 'Outputs'
   Bar "Bar_1" at 64,144 size 80x230; MinimumValue 0
      ProcessValue <- "Counter value"
   Bar "Bar_2" at 638,144 size 80x230; MinimumValue 0; MaximumValue 100
      ProcessValue <- "Assembled part counter value"
   TextField "Text field_4" at 610,101 size 156x23; Text 'Assembled Parts'
   IOField "I/O field_1" at 476,330 size 69x32; FormatPattern 999
      ProcessValue <- "Assembled part counter value"
   TextField "Text field_5" at 462,103 size 95x23; Text 'Metal peg'
   TextField "Text field_6" at 457,203 size 108x23; Text 'Plastic ring'
   IOField "I/O field_2" at 475,242 size 69x32; FormatPattern 999
      ProcessValue <- "Plastic ring counter value"
   IOField "I/O field_3" at 474,148 size 69x32; FormatPattern 999
      ProcessValue <- "Metal peg counter value"
   TextField "Text field_7" at 443,301 size 156x23; Text 'Assembled Parts'
   TextField "Text field_8" at 250,132 size 95x23; Text 'Metal peg'
   TextField "Text field_9" at 244,259 size 108x23; Text 'Plastic ring'
   IOField "I/O field_4" at 262,298 size 69x32; FormatPattern 999
      ProcessValue <- "Input plastic ring counter value"
   IOField "I/O field_5" at 262,177 size 69x32; FormatPattern 999
      ProcessValue <- "Input metal peg counter value"

screen "Temperature Control" 800x480, template "Template_1"
   TextField "HmiScreenItemData" at 80,196 size 640x25; Text 'Temperature Control'
   Button "Back" at 1,1 size 159x47; TextOff 'Back'
      on Release: ActivateScreen("Sorting Station Overview", 0)

screen "Alarm" 800x480, template "Template_1"
   TextField "HmiScreenItemData" at 80,196 size 640x25; Text 'Alarm'
   Button "Back" at 1,1 size 159x47; TextOff 'Back'
      on Release: ActivateScreen("Sorting Station Overview", 0)

screen "Exercise" 800x480, template "Template_1"
   TextField "HmiScreenItemData" at 80,196 size 640x25; Text 'Exercise'
   Button "Back" at 1,1 size 159x47; TextOff 'Back'
      on Release: ActivateScreen("Sorting Station Overview", 0)

screen "System screens" 800x480, template "Template_1"
   Button "Back" at 1,1 size 159x47; TextOff 'Back'
      on Release: ActivateScreen("Sorting Station Overview", 0)
   Button "HmiScreenItemData" at 36,95 size 159x47; TextOff 'SIMATIC PLC system diagnos...'; PictureOff "Navigates to SIMATIC PLC system diagnostics for TP700 Comfort 15.1.0.0"; PictureOn "Navigates to SIMATIC PLC system diagnostics for TP700 Comfort 15.1.0.0"
      on Release: ActivateScreen("SIMATIC PLC system diagnostics", 0)

screen "SIMATIC PLC system diagnostics" 800x480, template "Template_1"
   SysDiagControl "HmiScreenItemData" at 1,49 size 796x364
   Button "Back" at 1,1 size 159x47; TextOff 'Back'
      on Release: ActivateScreen("System screens", 0)
*)